REGION Network 3: Purga Bellis
   RUNG wire#powerrail
      Contact( "MC003" )
      Contact( "DB-PurgaComAlta".Habil_PurgaBellis )
      I_Contact( "Tag_55" )
      S_ODT(T_NO := "Tag_17", R := wire#w1, TV := #Aux1_MC003, BI =>, RET_VAL =>)
      wire#w2
      Coil( "MC003_EVP" )
   END_RUNG
   RUNG wire#powerrail
      I_Contact( "DB-PurgaComAlta".Habil_PurgaBellis )
   END_RUNG wire#w1
   RUNG wire#powerrail
      Contact( "DB-PurgaComAlta".Prueba_PurgaBellis )
      wire#w3
      I_Contact( "Tag_55" )
   END_RUNG wire#w2
   RUNG wire#powerrail
      Contact( "MC003_EVP" )
   END_RUNG wire#w3
   RUNG wire#w2
      S_ODT(T_NO := "Tag_55", TV := #Aux2_MC003, R :=, BI =>, RET_VAL =>)
   END_RUNG
   // the same network as SCL:
   #_s5time1 := S_ODT(T_NO := "Tag_17",
                      S := "MC003" AND "DB-PurgaComAlta".Habil_PurgaBellis AND NOT "Tag_55",
                      R := NOT "DB-PurgaComAlta".Habil_PurgaBellis,
                      TV := #Aux1_MC003,
                      Q => #_w1);
   "MC003_EVP" := #_w1 OR (("DB-PurgaComAlta".Prueba_PurgaBellis OR "MC003_EVP") AND NOT "Tag_55");
   #_s5time2 := S_ODT(T_NO := "Tag_55", S := "MC003_EVP", TV := #Aux2_MC003);
END_REGION

REGION Network 4
   RUNG wire#powerrail
      { S7_Templates := "SrcType := Int"; S7_GenerateENO := "TRUE" } Mul(in1 := "DB-PurgaComAlta".Toff_PurgaABC2, in2 := 6, out => #Aux1_MC001)
      { S7_Templates := "[SrcType := Int, DestType := Bcd16]"; S7_GenerateENO := "TRUE" } Convert(in := #Aux1_MC001, out => #Aux1_MC001)
      { S7_Templates := "SrcType := Int"; S7_GenerateENO := "TRUE" } Add(in1 := #Aux1_MC001, in2 := 16#3000, out => #Aux1_MC001)
   END_RUNG
   // the same network as SCL:
   // ENO of a box is taken as its EN; it also drops when the box reports an error
   #Aux1_MC001 := "DB-PurgaComAlta".Toff_PurgaABC2 * 6;
   #Aux1_MC001 := INT_TO_BCD16(#Aux1_MC001);
   #Aux1_MC001 := #Aux1_MC001 + 16#3000;
END_REGION

REGION Network 5
   RUNG wire#powerrail
      { S7_Templates := "SrcType := Int"; S7_GenerateENO := "TRUE" } Mul(in1 := "DB-PurgaComAlta".Ton_PurgaABC2, in2 := 10, out => #Aux2_MC001)
      { S7_Templates := "[SrcType := Int, DestType := Bcd16]"; S7_GenerateENO := "TRUE" } Convert(in := #Aux2_MC001, out => #Aux2_MC001)
      { S7_Templates := "SrcType := Int"; S7_GenerateENO := "TRUE" } Add(in1 := #Aux2_MC001, in2 := 16#1000, out => #Aux2_MC001)
   END_RUNG
   // the same network as SCL:
   // ENO of a box is taken as its EN; it also drops when the box reports an error
   #Aux2_MC001 := "DB-PurgaComAlta".Ton_PurgaABC2 * 10;
   #Aux2_MC001 := INT_TO_BCD16(#Aux2_MC001);
   #Aux2_MC001 := #Aux2_MC001 + 16#1000;
END_REGION

REGION Network 6: Purga ABC2
   RUNG wire#powerrail
      Contact( "MC001" )
      Contact( "DB-PurgaComAlta".Habil_PurgaABC2 )
      I_Contact( "Tag_65" )
      S_ODT(T_NO := "Tag_64", R := wire#w1, TV := #Aux1_MC001, BI =>, RET_VAL =>)
      I_Contact( "MC003_EVP" )
      wire#w2
      Coil( "MC001_EVP" )
   END_RUNG
   RUNG wire#powerrail
      I_Contact( "DB-PurgaComAlta".Habil_PurgaABC2 )
   END_RUNG wire#w1
   RUNG wire#powerrail
      Contact( "DB-PurgaComAlta".Prueba_PurgaABC2 )
      wire#w3
      I_Contact( "Tag_65" )
   END_RUNG wire#w2
   RUNG wire#powerrail
      Contact( "MC001_EVP" )
   END_RUNG wire#w3
   RUNG wire#w2
      S_ODT(T_NO := "Tag_65", TV := #Aux2_MC001, R :=, BI =>, RET_VAL =>)
   END_RUNG
   // the same network as SCL:
   #_s5time1 := S_ODT(T_NO := "Tag_64",
                      S := "MC001" AND "DB-PurgaComAlta".Habil_PurgaABC2 AND NOT "Tag_65",
                      R := NOT "DB-PurgaComAlta".Habil_PurgaABC2,
                      TV := #Aux1_MC001,
                      Q => #_w1);
   "MC001_EVP" := (#_w1 AND NOT "MC003_EVP") OR (("DB-PurgaComAlta".Prueba_PurgaABC2 OR "MC001_EVP") AND NOT "Tag_65");
   #_s5time2 := S_ODT(T_NO := "Tag_65", S := "MC001_EVP", TV := #Aux2_MC001);
END_REGION

REGION Network 7
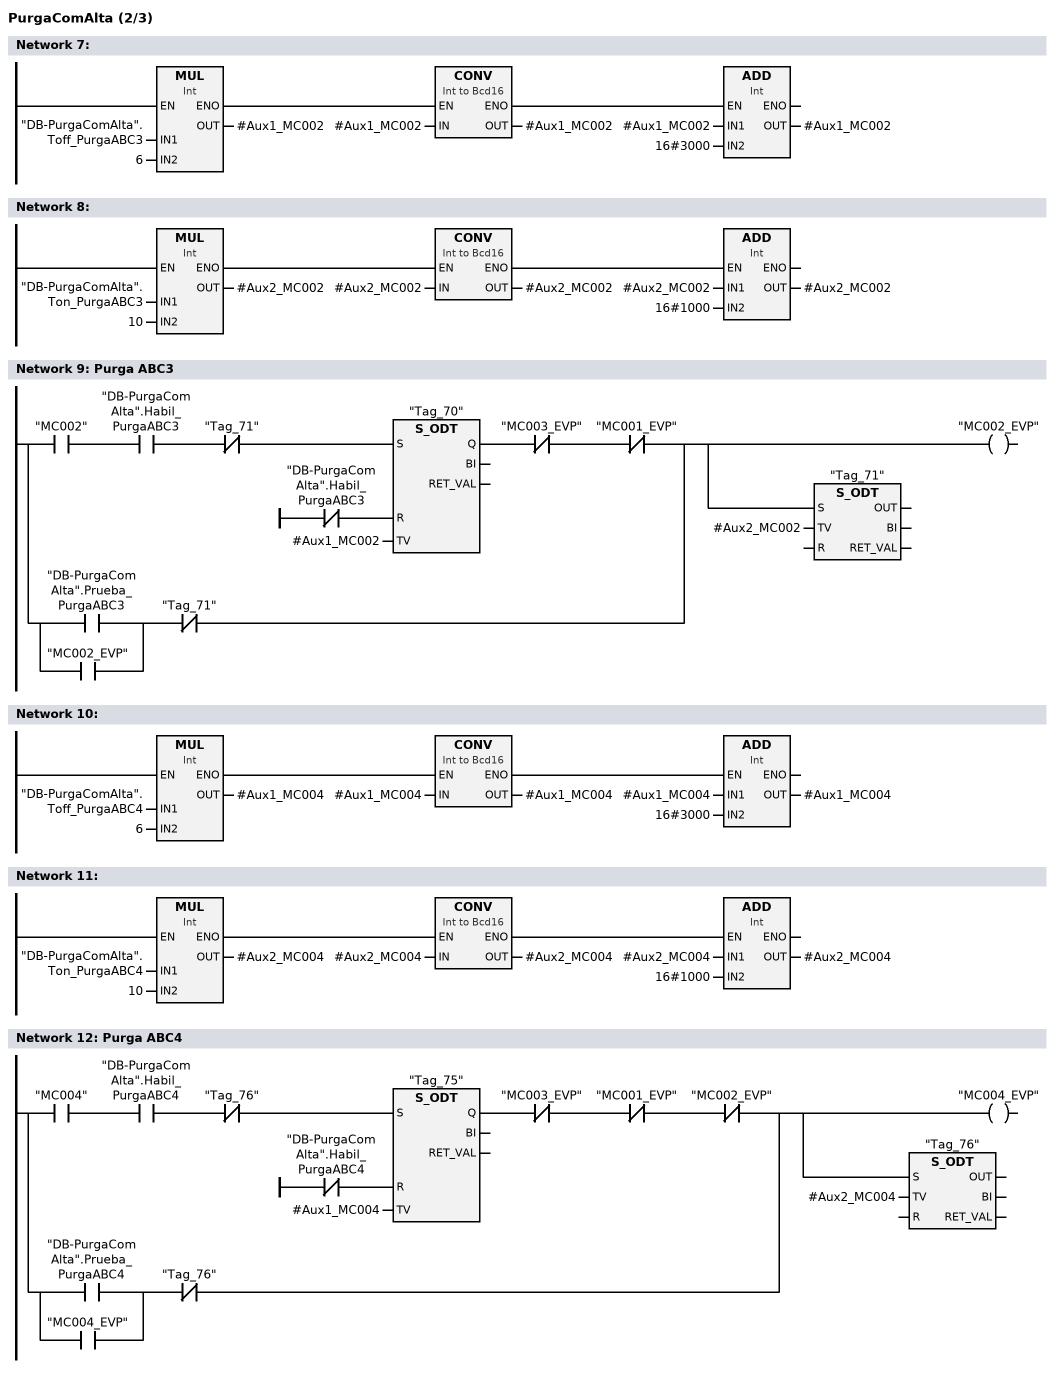
   RUNG wire#powerrail
      { S7_Templates := "SrcType := Int"; S7_GenerateENO := "TRUE" } Mul(in1 := "DB-PurgaComAlta".Toff_PurgaABC3, in2 := 6, out => #Aux1_MC002)
      { S7_Templates := "[SrcType := Int, DestType := Bcd16]"; S7_GenerateENO := "TRUE" } Convert(in := #Aux1_MC002, out => #Aux1_MC002)
      { S7_Templates := "SrcType := Int"; S7_GenerateENO := "TRUE" } Add(in1 := #Aux1_MC002, in2 := 16#3000, out => #Aux1_MC002)
   END_RUNG
   // the same network as SCL:
   // ENO of a box is taken as its EN; it also drops when the box reports an error
   #Aux1_MC002 := "DB-PurgaComAlta".Toff_PurgaABC3 * 6;
   #Aux1_MC002 := INT_TO_BCD16(#Aux1_MC002);
   #Aux1_MC002 := #Aux1_MC002 + 16#3000;
END_REGION

REGION Network 8
   RUNG wire#powerrail
      { S7_Templates := "SrcType := Int"; S7_GenerateENO := "TRUE" } Mul(in1 := "DB-PurgaComAlta".Ton_PurgaABC3, in2 := 10, out => #Aux2_MC002)
      { S7_Templates := "[SrcType := Int, DestType := Bcd16]"; S7_GenerateENO := "TRUE" } Convert(in := #Aux2_MC002, out => #Aux2_MC002)
      { S7_Templates := "SrcType := Int"; S7_GenerateENO := "TRUE" } Add(in1 := #Aux2_MC002, in2 := 16#1000, out => #Aux2_MC002)
   END_RUNG
   // the same network as SCL:
   // ENO of a box is taken as its EN; it also drops when the box reports an error
   #Aux2_MC002 := "DB-PurgaComAlta".Ton_PurgaABC3 * 10;
   #Aux2_MC002 := INT_TO_BCD16(#Aux2_MC002);
   #Aux2_MC002 := #Aux2_MC002 + 16#1000;
END_REGION

REGION Network 9: Purga ABC3
   RUNG wire#powerrail
      Contact( "MC002" )
      Contact( "DB-PurgaComAlta".Habil_PurgaABC3 )
      I_Contact( "Tag_71" )
      S_ODT(T_NO := "Tag_70", R := wire#w1, TV := #Aux1_MC002, BI =>, RET_VAL =>)
      I_Contact( "MC003_EVP" )
      I_Contact( "MC001_EVP" )
      wire#w2
      Coil( "MC002_EVP" )
   END_RUNG
   RUNG wire#powerrail
      I_Contact( "DB-PurgaComAlta".Habil_PurgaABC3 )
   END_RUNG wire#w1
   RUNG wire#powerrail
      Contact( "DB-PurgaComAlta".Prueba_PurgaABC3 )
      wire#w3
      I_Contact( "Tag_71" )
   END_RUNG wire#w2
   RUNG wire#powerrail
      Contact( "MC002_EVP" )
   END_RUNG wire#w3
   RUNG wire#w2
      S_ODT(T_NO := "Tag_71", TV := #Aux2_MC002, R :=, BI =>, RET_VAL =>)
   END_RUNG
   // the same network as SCL:
   #_s5time1 := S_ODT(T_NO := "Tag_70",
                      S := "MC002" AND "DB-PurgaComAlta".Habil_PurgaABC3 AND NOT "Tag_71",
                      R := NOT "DB-PurgaComAlta".Habil_PurgaABC3,
                      TV := #Aux1_MC002,
                      Q => #_w1);
   "MC002_EVP" := (#_w1 AND NOT "MC003_EVP" AND NOT "MC001_EVP") OR (("DB-PurgaComAlta".Prueba_PurgaABC3 OR "MC002_EVP") AND NOT "Tag_71");
   #_s5time2 := S_ODT(T_NO := "Tag_71", S := "MC002_EVP", TV := #Aux2_MC002);
END_REGION

REGION Network 10
   RUNG wire#powerrail
      { S7_Templates := "SrcType := Int"; S7_GenerateENO := "TRUE" } Mul(in1 := "DB-PurgaComAlta".Toff_PurgaABC4, in2 := 6, out => #Aux1_MC004)
      { S7_Templates := "[SrcType := Int, DestType := Bcd16]"; S7_GenerateENO := "TRUE" } Convert(in := #Aux1_MC004, out => #Aux1_MC004)
      { S7_Templates := "SrcType := Int"; S7_GenerateENO := "TRUE" } Add(in1 := #Aux1_MC004, in2 := 16#3000, out => #Aux1_MC004)
   END_RUNG
   // the same network as SCL:
   // ENO of a box is taken as its EN; it also drops when the box reports an error
   #Aux1_MC004 := "DB-PurgaComAlta".Toff_PurgaABC4 * 6;
   #Aux1_MC004 := INT_TO_BCD16(#Aux1_MC004);
   #Aux1_MC004 := #Aux1_MC004 + 16#3000;
END_REGION

REGION Network 11
   RUNG wire#powerrail
      { S7_Templates := "SrcType := Int"; S7_GenerateENO := "TRUE" } Mul(in1 := "DB-PurgaComAlta".Ton_PurgaABC4, in2 := 10, out => #Aux2_MC004)
      { S7_Templates := "[SrcType := Int, DestType := Bcd16]"; S7_GenerateENO := "TRUE" } Convert(in := #Aux2_MC004, out => #Aux2_MC004)
      { S7_Templates := "SrcType := Int"; S7_GenerateENO := "TRUE" } Add(in1 := #Aux2_MC004, in2 := 16#1000, out => #Aux2_MC004)
   END_RUNG
   // the same network as SCL:
   // ENO of a box is taken as its EN; it also drops when the box reports an error
   #Aux2_MC004 := "DB-PurgaComAlta".Ton_PurgaABC4 * 10;
   #Aux2_MC004 := INT_TO_BCD16(#Aux2_MC004);
   #Aux2_MC004 := #Aux2_MC004 + 16#1000;
END_REGION

REGION Network 12: Purga ABC4
   RUNG wire#powerrail
      Contact( "MC004" )
      Contact( "DB-PurgaComAlta".Habil_PurgaABC4 )
      I_Contact( "Tag_76" )
      S_ODT(T_NO := "Tag_75", R := wire#w1, TV := #Aux1_MC004, BI =>, RET_VAL =>)
      I_Contact( "MC003_EVP" )
      I_Contact( "MC001_EVP" )
      I_Contact( "MC002_EVP" )
      wire#w2
      Coil( "MC004_EVP" )
   END_RUNG
   RUNG wire#powerrail
      I_Contact( "DB-PurgaComAlta".Habil_PurgaABC4 )
   END_RUNG wire#w1
   RUNG wire#powerrail
      Contact( "DB-PurgaComAlta".Prueba_PurgaABC4 )
      wire#w3
      I_Contact( "Tag_76" )
   END_RUNG wire#w2
   RUNG wire#powerrail
      Contact( "MC004_EVP" )
   END_RUNG wire#w3
   RUNG wire#w2
      S_ODT(T_NO := "Tag_76", TV := #Aux2_MC004, R :=, BI =>, RET_VAL =>)
   END_RUNG
   // the same network as SCL:
   #_s5time1 := S_ODT(T_NO := "Tag_75",
                      S := "MC004" AND "DB-PurgaComAlta".Habil_PurgaABC4 AND NOT "Tag_76",
                      R := NOT "DB-PurgaComAlta".Habil_PurgaABC4,
                      TV := #Aux1_MC004,
                      Q => #_w1);
   "MC004_EVP" := (#_w1 AND NOT "MC003_EVP" AND NOT "MC001_EVP" AND NOT "MC002_EVP") OR (("DB-PurgaComAlta".Prueba_PurgaABC4 OR "MC004_EVP") AND NOT "Tag_76");
   #_s5time2 := S_ODT(T_NO := "Tag_76", S := "MC004_EVP", TV := #Aux2_MC004);
END_REGION

REGION Network 13
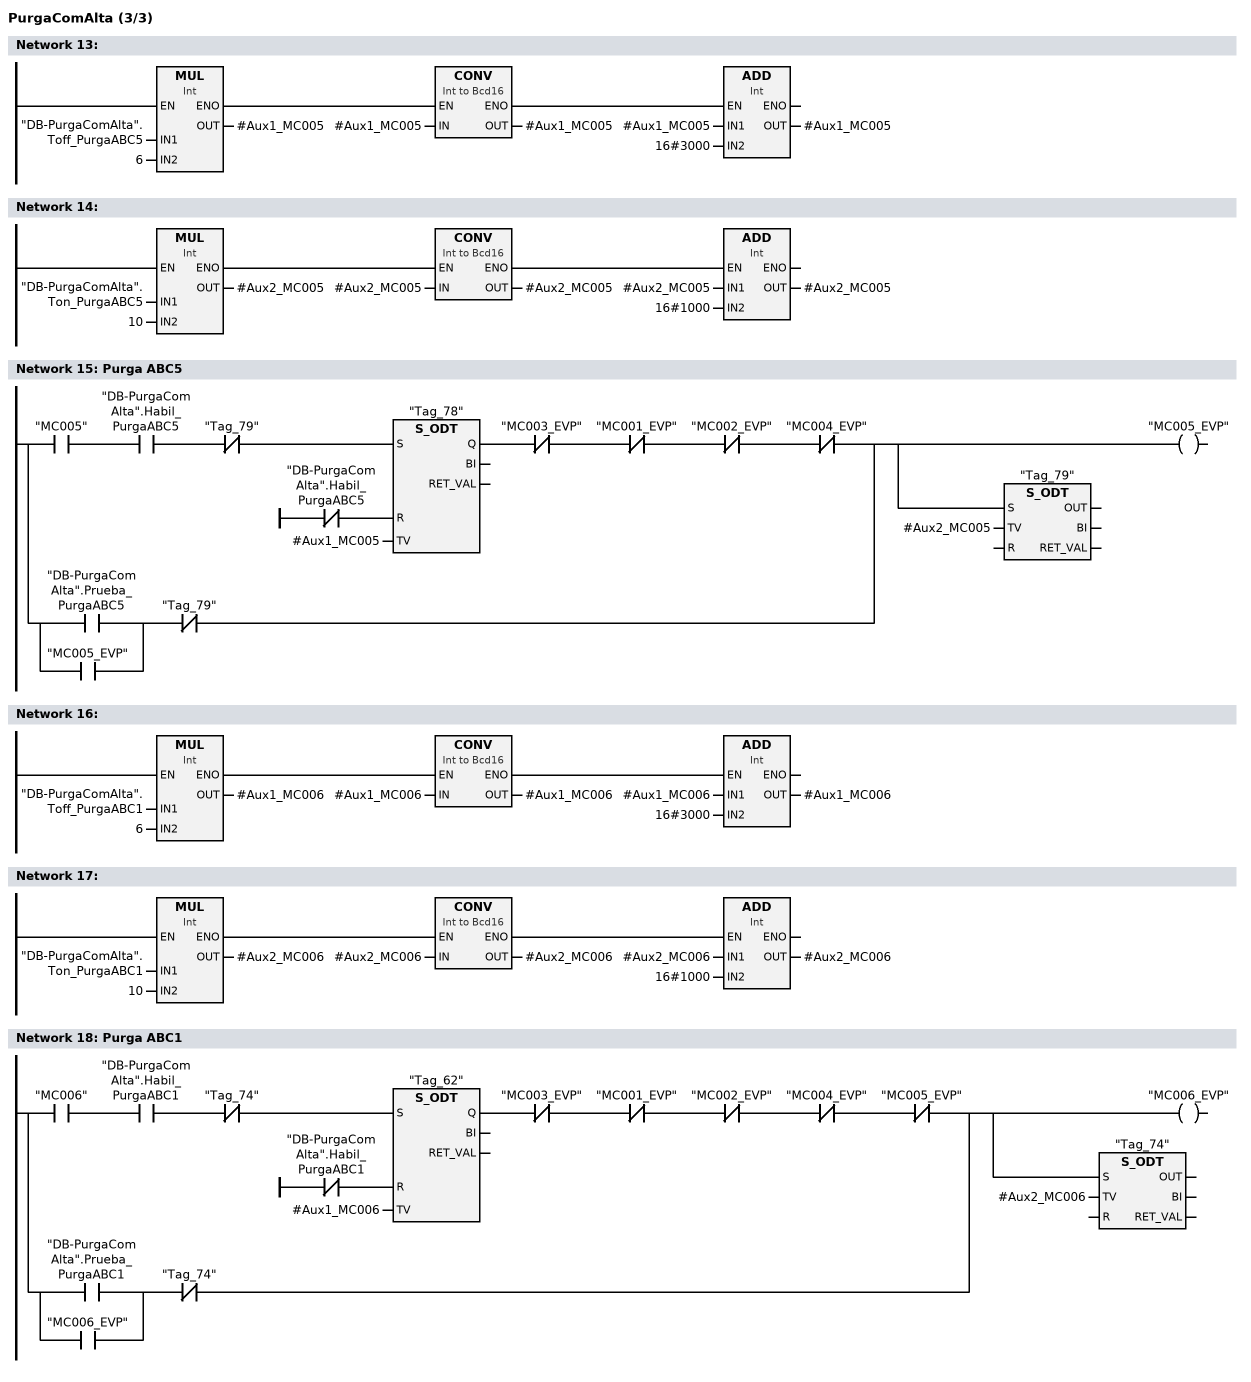
   RUNG wire#powerrail
      { S7_Templates := "SrcType := Int"; S7_GenerateENO := "TRUE" } Mul(in1 := "DB-PurgaComAlta".Toff_PurgaABC5, in2 := 6, out => #Aux1_MC005)
      { S7_Templates := "[SrcType := Int, DestType := Bcd16]"; S7_GenerateENO := "TRUE" } Convert(in := #Aux1_MC005, out => #Aux1_MC005)
      { S7_Templates := "SrcType := Int"; S7_GenerateENO := "TRUE" } Add(in1 := #Aux1_MC005, in2 := 16#3000, out => #Aux1_MC005)
   END_RUNG
   // the same network as SCL:
   // ENO of a box is taken as its EN; it also drops when the box reports an error
   #Aux1_MC005 := "DB-PurgaComAlta".Toff_PurgaABC5 * 6;
   #Aux1_MC005 := INT_TO_BCD16(#Aux1_MC005);
   #Aux1_MC005 := #Aux1_MC005 + 16#3000;
END_REGION

REGION Network 14
   RUNG wire#powerrail
      { S7_Templates := "SrcType := Int"; S7_GenerateENO := "TRUE" } Mul(in1 := "DB-PurgaComAlta".Ton_PurgaABC5, in2 := 10, out => #Aux2_MC005)
      { S7_Templates := "[SrcType := Int, DestType := Bcd16]"; S7_GenerateENO := "TRUE" } Convert(in := #Aux2_MC005, out => #Aux2_MC005)
      { S7_Templates := "SrcType := Int"; S7_GenerateENO := "TRUE" } Add(in1 := #Aux2_MC005, in2 := 16#1000, out => #Aux2_MC005)
   END_RUNG
   // the same network as SCL:
   // ENO of a box is taken as its EN; it also drops when the box reports an error
   #Aux2_MC005 := "DB-PurgaComAlta".Ton_PurgaABC5 * 10;
   #Aux2_MC005 := INT_TO_BCD16(#Aux2_MC005);
   #Aux2_MC005 := #Aux2_MC005 + 16#1000;
END_REGION

REGION Network 15: Purga ABC5
   RUNG wire#powerrail
      Contact( "MC005" )
      Contact( "DB-PurgaComAlta".Habil_PurgaABC5 )
      I_Contact( "Tag_79" )
      S_ODT(T_NO := "Tag_78", R := wire#w1, TV := #Aux1_MC005, BI =>, RET_VAL =>)
      I_Contact( "MC003_EVP" )
      I_Contact( "MC001_EVP" )
      I_Contact( "MC002_EVP" )
      I_Contact( "MC004_EVP" )
      wire#w2
      Coil( "MC005_EVP" )
   END_RUNG
   RUNG wire#powerrail
      I_Contact( "DB-PurgaComAlta".Habil_PurgaABC5 )
   END_RUNG wire#w1
   RUNG wire#powerrail
      Contact( "DB-PurgaComAlta".Prueba_PurgaABC5 )
      wire#w3
      I_Contact( "Tag_79" )
   END_RUNG wire#w2
   RUNG wire#powerrail
      Contact( "MC005_EVP" )
   END_RUNG wire#w3
   RUNG wire#w2
      S_ODT(T_NO := "Tag_79", TV := #Aux2_MC005, R :=, BI =>, RET_VAL =>)
   END_RUNG
   // the same network as SCL:
   #_s5time1 := S_ODT(T_NO := "Tag_78",
                      S := "MC005" AND "DB-PurgaComAlta".Habil_PurgaABC5 AND NOT "Tag_79",
                      R := NOT "DB-PurgaComAlta".Habil_PurgaABC5,
                      TV := #Aux1_MC005,
                      Q => #_w1);
   "MC005_EVP" := (#_w1 AND NOT "MC003_EVP" AND NOT "MC001_EVP" AND NOT "MC002_EVP" AND NOT "MC004_EVP") OR (("DB-PurgaComAlta".Prueba_PurgaABC5 OR "MC005_EVP") AND NOT "Tag_79");
   #_s5time2 := S_ODT(T_NO := "Tag_79", S := "MC005_EVP", TV := #Aux2_MC005);
END_REGION

REGION Network 16
   RUNG wire#powerrail
      { S7_Templates := "SrcType := Int"; S7_GenerateENO := "TRUE" } Mul(in1 := "DB-PurgaComAlta".Toff_PurgaABC1, in2 := 6, out => #Aux1_MC006)
      { S7_Templates := "[SrcType := Int, DestType := Bcd16]"; S7_GenerateENO := "TRUE" } Convert(in := #Aux1_MC006, out => #Aux1_MC006)
      { S7_Templates := "SrcType := Int"; S7_GenerateENO := "TRUE" } Add(in1 := #Aux1_MC006, in2 := 16#3000, out => #Aux1_MC006)
   END_RUNG
   // the same network as SCL:
   // ENO of a box is taken as its EN; it also drops when the box reports an error
   #Aux1_MC006 := "DB-PurgaComAlta".Toff_PurgaABC1 * 6;
   #Aux1_MC006 := INT_TO_BCD16(#Aux1_MC006);
   #Aux1_MC006 := #Aux1_MC006 + 16#3000;
END_REGION

REGION Network 17
   RUNG wire#powerrail
      { S7_Templates := "SrcType := Int"; S7_GenerateENO := "TRUE" } Mul(in1 := "DB-PurgaComAlta".Ton_PurgaABC1, in2 := 10, out => #Aux2_MC006)
      { S7_Templates := "[SrcType := Int, DestType := Bcd16]"; S7_GenerateENO := "TRUE" } Convert(in := #Aux2_MC006, out => #Aux2_MC006)
      { S7_Templates := "SrcType := Int"; S7_GenerateENO := "TRUE" } Add(in1 := #Aux2_MC006, in2 := 16#1000, out => #Aux2_MC006)
   END_RUNG
   // the same network as SCL:
   // ENO of a box is taken as its EN; it also drops when the box reports an error
   #Aux2_MC006 := "DB-PurgaComAlta".Ton_PurgaABC1 * 10;
   #Aux2_MC006 := INT_TO_BCD16(#Aux2_MC006);
   #Aux2_MC006 := #Aux2_MC006 + 16#1000;
END_REGION

REGION Network 18: Purga ABC1
   RUNG wire#powerrail
      Contact( "MC006" )
      Contact( "DB-PurgaComAlta".Habil_PurgaABC1 )
      I_Contact( "Tag_74" )
      S_ODT(T_NO := "Tag_62", R := wire#w1, TV := #Aux1_MC006, BI =>, RET_VAL =>)
      I_Contact( "MC003_EVP" )
      I_Contact( "MC001_EVP" )
      I_Contact( "MC002_EVP" )
      I_Contact( "MC004_EVP" )
      I_Contact( "MC005_EVP" )
      wire#w2
      Coil( "MC006_EVP" )
   END_RUNG
   RUNG wire#powerrail
      I_Contact( "DB-PurgaComAlta".Habil_PurgaABC1 )
   END_RUNG wire#w1
   RUNG wire#powerrail
      Contact( "DB-PurgaComAlta".Prueba_PurgaABC1 )
      wire#w3
      I_Contact( "Tag_74" )
   END_RUNG wire#w2
   RUNG wire#powerrail
      Contact( "MC006_EVP" )
   END_RUNG wire#w3
   RUNG wire#w2
      S_ODT(T_NO := "Tag_74", TV := #Aux2_MC006, R :=, BI =>, RET_VAL =>)
   END_RUNG
   // the same network as SCL:
   #_s5time1 := S_ODT(T_NO := "Tag_62",
                      S := "MC006" AND "DB-PurgaComAlta".Habil_PurgaABC1 AND NOT "Tag_74",
                      R := NOT "DB-PurgaComAlta".Habil_PurgaABC1,
                      TV := #Aux1_MC006,
                      Q => #_w1);
   "MC006_EVP" := (#_w1 AND NOT "MC003_EVP" AND NOT "MC001_EVP" AND NOT "MC002_EVP" AND NOT "MC004_EVP" AND NOT "MC005_EVP") OR (("DB-PurgaComAlta".Prueba_PurgaABC1 OR "MC006_EVP") AND NOT "Tag_74");
   #_s5time2 := S_ODT(T_NO := "Tag_74", S := "MC006_EVP", TV := #Aux2_MC006);
END_REGION
END_FUNCTION

// folder: Compresores/Alta/Máquina de Estados

FUNCTION "LogMaqEstGeneral" : Void   // FC35, LAD
{ S7_Optimized_Access := 'FALSE' }
VERSION : 0.1
   VAR_TEMP
      Temp_0 : Bool;
      Temp_1 : Bool;
      Temp_2 : Bool;
      Temp_3 : Bool;
      Temp_4 : Bool;
      Temp_5 : Bool;
      Temp_6 : Bool;
      Temp_7 : Bool;
      Temp_8 : Bool;
      Temp_9 : Bool;
      Temp_10 : Bool;
      Temp_11 : Bool;
   END_VAR
BEGIN

REGION Network 1
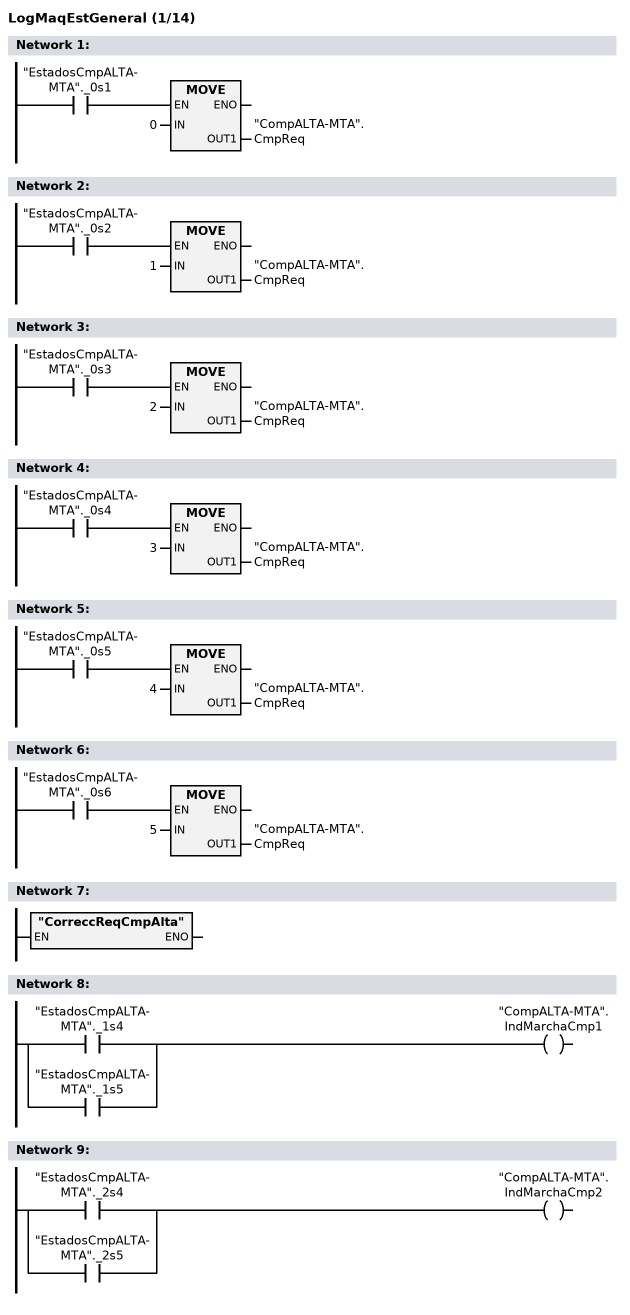
   RUNG wire#powerrail
      Contact( "EstadosCmpALTA-MTA"._0s1 )
      { S7_GenerateENO := "TRUE" } Move(in := 0, out1 => "CompALTA-MTA".CmpReq)
   END_RUNG
   // the same network as SCL:
   IF "EstadosCmpALTA-MTA"._0s1 THEN "CompALTA-MTA".CmpReq := 0; END_IF;
END_REGION

REGION Network 2
   RUNG wire#powerrail
      Contact( "EstadosCmpALTA-MTA"._0s2 )
      { S7_GenerateENO := "TRUE" } Move(in := 1, out1 => "CompALTA-MTA".CmpReq)
   END_RUNG
   // the same network as SCL:
   IF "EstadosCmpALTA-MTA"._0s2 THEN "CompALTA-MTA".CmpReq := 1; END_IF;
END_REGION

REGION Network 3
   RUNG wire#powerrail
      Contact( "EstadosCmpALTA-MTA"._0s3 )
      { S7_GenerateENO := "TRUE" } Move(in := 2, out1 => "CompALTA-MTA".CmpReq)
   END_RUNG
   // the same network as SCL:
   IF "EstadosCmpALTA-MTA"._0s3 THEN "CompALTA-MTA".CmpReq := 2; END_IF;
END_REGION

REGION Network 4
   RUNG wire#powerrail
      Contact( "EstadosCmpALTA-MTA"._0s4 )
      { S7_GenerateENO := "TRUE" } Move(in := 3, out1 => "CompALTA-MTA".CmpReq)
   END_RUNG
   // the same network as SCL:
   IF "EstadosCmpALTA-MTA"._0s4 THEN "CompALTA-MTA".CmpReq := 3; END_IF;
END_REGION

REGION Network 5
   RUNG wire#powerrail
      Contact( "EstadosCmpALTA-MTA"._0s5 )
      { S7_GenerateENO := "TRUE" } Move(in := 4, out1 => "CompALTA-MTA".CmpReq)
   END_RUNG
   // the same network as SCL:
   IF "EstadosCmpALTA-MTA"._0s5 THEN "CompALTA-MTA".CmpReq := 4; END_IF;
END_REGION

REGION Network 6
   RUNG wire#powerrail
      Contact( "EstadosCmpALTA-MTA"._0s6 )
      { S7_GenerateENO := "TRUE" } Move(in := 5, out1 => "CompALTA-MTA".CmpReq)
   END_RUNG
   // the same network as SCL:
   IF "EstadosCmpALTA-MTA"._0s6 THEN "CompALTA-MTA".CmpReq := 5; END_IF;
END_REGION

REGION Network 7
   RUNG wire#powerrail
      "CorreccReqCmpAlta"()
   END_RUNG
   // the same network as SCL:
   "CorreccReqCmpAlta"();
END_REGION

REGION Network 8
   RUNG wire#powerrail
      Contact( "EstadosCmpALTA-MTA"._1s4 )
      wire#w1
      Coil( "CompALTA-MTA".IndMarchaCmp1 )
   END_RUNG
   RUNG wire#powerrail
      Contact( "EstadosCmpALTA-MTA"._1s5 )
   END_RUNG wire#w1
   // the same network as SCL:
   "CompALTA-MTA".IndMarchaCmp1 := "EstadosCmpALTA-MTA"._1s4 OR "EstadosCmpALTA-MTA"._1s5;
END_REGION

REGION Network 9
   RUNG wire#powerrail
      Contact( "EstadosCmpALTA-MTA"._2s4 )
      wire#w1
      Coil( "CompALTA-MTA".IndMarchaCmp2 )
   END_RUNG
   RUNG wire#powerrail
      Contact( "EstadosCmpALTA-MTA"._2s5 )
   END_RUNG wire#w1
   // the same network as SCL:
   "CompALTA-MTA".IndMarchaCmp2 := "EstadosCmpALTA-MTA"._2s4 OR "EstadosCmpALTA-MTA"._2s5;
END_REGION

REGION Network 10
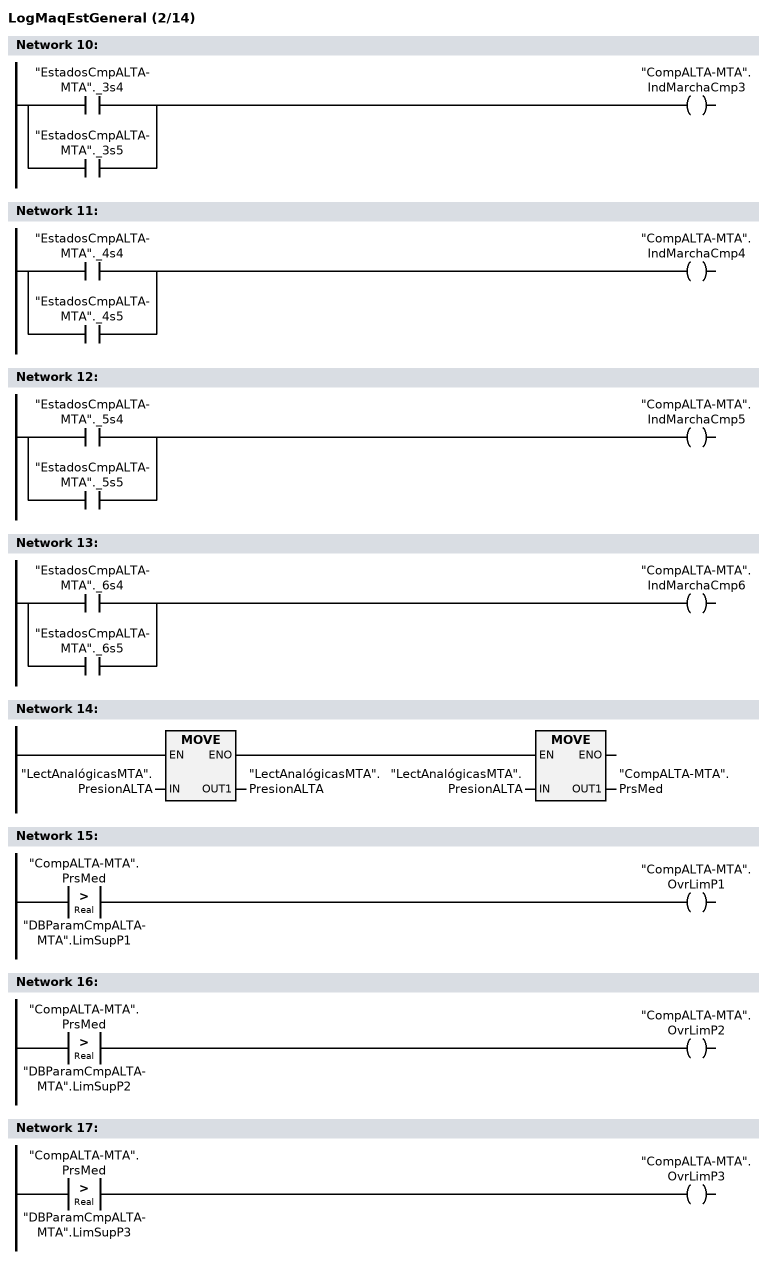
   RUNG wire#powerrail
      Contact( "EstadosCmpALTA-MTA"._3s4 )
      wire#w1
      Coil( "CompALTA-MTA".IndMarchaCmp3 )
   END_RUNG
   RUNG wire#powerrail
      Contact( "EstadosCmpALTA-MTA"._3s5 )
   END_RUNG wire#w1
   // the same network as SCL:
   "CompALTA-MTA".IndMarchaCmp3 := "EstadosCmpALTA-MTA"._3s4 OR "EstadosCmpALTA-MTA"._3s5;
END_REGION

REGION Network 11
   RUNG wire#powerrail
      Contact( "EstadosCmpALTA-MTA"._4s4 )
      wire#w1
      Coil( "CompALTA-MTA".IndMarchaCmp4 )
   END_RUNG
   RUNG wire#powerrail
      Contact( "EstadosCmpALTA-MTA"._4s5 )
   END_RUNG wire#w1
   // the same network as SCL:
   "CompALTA-MTA".IndMarchaCmp4 := "EstadosCmpALTA-MTA"._4s4 OR "EstadosCmpALTA-MTA"._4s5;
END_REGION

REGION Network 12
   RUNG wire#powerrail
      Contact( "EstadosCmpALTA-MTA"._5s4 )
      wire#w1
      Coil( "CompALTA-MTA".IndMarchaCmp5 )
   END_RUNG
   RUNG wire#powerrail
      Contact( "EstadosCmpALTA-MTA"._5s5 )
   END_RUNG wire#w1
   // the same network as SCL:
   "CompALTA-MTA".IndMarchaCmp5 := "EstadosCmpALTA-MTA"._5s4 OR "EstadosCmpALTA-MTA"._5s5;
END_REGION

REGION Network 13
   RUNG wire#powerrail
      Contact( "EstadosCmpALTA-MTA"._6s4 )
      wire#w1
      Coil( "CompALTA-MTA".IndMarchaCmp6 )
   END_RUNG
   RUNG wire#powerrail
      Contact( "EstadosCmpALTA-MTA"._6s5 )
   END_RUNG wire#w1
   // the same network as SCL:
   "CompALTA-MTA".IndMarchaCmp6 := "EstadosCmpALTA-MTA"._6s4 OR "EstadosCmpALTA-MTA"._6s5;
END_REGION

REGION Network 14
   RUNG wire#powerrail
      { S7_GenerateENO := "TRUE" } Move(in := "LectAnalógicasMTA".PresionALTA, out1 => "LectAnalógicasMTA".PresionALTA)
      { S7_GenerateENO := "TRUE" } Move(in := "LectAnalógicasMTA".PresionALTA, out1 => "CompALTA-MTA".PrsMed)
   END_RUNG
   // the same network as SCL:
   // ENO of a box is taken as its EN; it also drops when the box reports an error
   "LectAnalógicasMTA".PresionALTA := "LectAnalógicasMTA".PresionALTA;
   "CompALTA-MTA".PrsMed := "LectAnalógicasMTA".PresionALTA;
END_REGION

REGION Network 15
   RUNG wire#powerrail
      { S7_Templates := "SrcType := Real" } GT_Contact(in1 := "CompALTA-MTA".PrsMed, in2 := "DBParamCmpALTA-MTA".LimSupP1)
      Coil( "CompALTA-MTA".OvrLimP1 )
   END_RUNG
   // the same network as SCL:
   "CompALTA-MTA".OvrLimP1 := "CompALTA-MTA".PrsMed > "DBParamCmpALTA-MTA".LimSupP1;
END_REGION

REGION Network 16
   RUNG wire#powerrail
      { S7_Templates := "SrcType := Real" } GT_Contact(in1 := "CompALTA-MTA".PrsMed, in2 := "DBParamCmpALTA-MTA".LimSupP2)
      Coil( "CompALTA-MTA".OvrLimP2 )
   END_RUNG
   // the same network as SCL:
   "CompALTA-MTA".OvrLimP2 := "CompALTA-MTA".PrsMed > "DBParamCmpALTA-MTA".LimSupP2;
END_REGION

REGION Network 17
   RUNG wire#powerrail
      { S7_Templates := "SrcType := Real" } GT_Contact(in1 := "CompALTA-MTA".PrsMed, in2 := "DBParamCmpALTA-MTA".LimSupP3)
      Coil( "CompALTA-MTA".OvrLimP3 )
   END_RUNG
   // the same network as SCL:
   "CompALTA-MTA".OvrLimP3 := "CompALTA-MTA".PrsMed > "DBParamCmpALTA-MTA".LimSupP3;
END_REGION

REGION Network 18
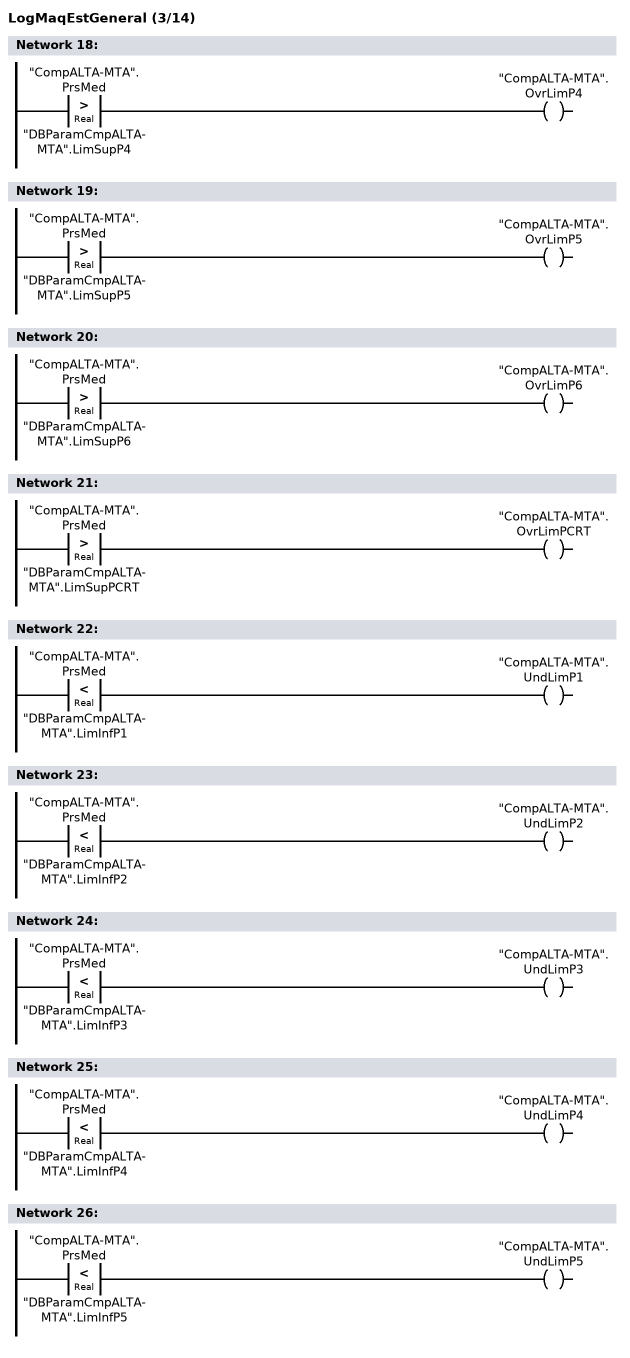
   RUNG wire#powerrail
      { S7_Templates := "SrcType := Real" } GT_Contact(in1 := "CompALTA-MTA".PrsMed, in2 := "DBParamCmpALTA-MTA".LimSupP4)
      Coil( "CompALTA-MTA".OvrLimP4 )
   END_RUNG
   // the same network as SCL:
   "CompALTA-MTA".OvrLimP4 := "CompALTA-MTA".PrsMed > "DBParamCmpALTA-MTA".LimSupP4;
END_REGION

REGION Network 19
   RUNG wire#powerrail
      { S7_Templates := "SrcType := Real" } GT_Contact(in1 := "CompALTA-MTA".PrsMed, in2 := "DBParamCmpALTA-MTA".LimSupP5)
      Coil( "CompALTA-MTA".OvrLimP5 )
   END_RUNG
   // the same network as SCL:
   "CompALTA-MTA".OvrLimP5 := "CompALTA-MTA".PrsMed > "DBParamCmpALTA-MTA".LimSupP5;
END_REGION

REGION Network 20
   RUNG wire#powerrail
      { S7_Templates := "SrcType := Real" } GT_Contact(in1 := "CompALTA-MTA".PrsMed, in2 := "DBParamCmpALTA-MTA".LimSupP6)
      Coil( "CompALTA-MTA".OvrLimP6 )
   END_RUNG
   // the same network as SCL:
   "CompALTA-MTA".OvrLimP6 := "CompALTA-MTA".PrsMed > "DBParamCmpALTA-MTA".LimSupP6;
END_REGION

REGION Network 21
   RUNG wire#powerrail
      { S7_Templates := "SrcType := Real" } GT_Contact(in1 := "CompALTA-MTA".PrsMed, in2 := "DBParamCmpALTA-MTA".LimSupPCRT)
      Coil( "CompALTA-MTA".OvrLimPCRT )
   END_RUNG
   // the same network as SCL:
   "CompALTA-MTA".OvrLimPCRT := "CompALTA-MTA".PrsMed > "DBParamCmpALTA-MTA".LimSupPCRT;
END_REGION

REGION Network 22
   RUNG wire#powerrail
      { S7_Templates := "SrcType := Real" } LT_Contact(in1 := "CompALTA-MTA".PrsMed, in2 := "DBParamCmpALTA-MTA".LimInfP1)
      Coil( "CompALTA-MTA".UndLimP1 )
   END_RUNG
   // the same network as SCL:
   "CompALTA-MTA".UndLimP1 := "CompALTA-MTA".PrsMed < "DBParamCmpALTA-MTA".LimInfP1;
END_REGION

REGION Network 23
   RUNG wire#powerrail
      { S7_Templates := "SrcType := Real" } LT_Contact(in1 := "CompALTA-MTA".PrsMed, in2 := "DBParamCmpALTA-MTA".LimInfP2)
      Coil( "CompALTA-MTA".UndLimP2 )
   END_RUNG
   // the same network as SCL:
   "CompALTA-MTA".UndLimP2 := "CompALTA-MTA".PrsMed < "DBParamCmpALTA-MTA".LimInfP2;
END_REGION

REGION Network 24
   RUNG wire#powerrail
      { S7_Templates := "SrcType := Real" } LT_Contact(in1 := "CompALTA-MTA".PrsMed, in2 := "DBParamCmpALTA-MTA".LimInfP3)
      Coil( "CompALTA-MTA".UndLimP3 )
   END_RUNG
   // the same network as SCL:
   "CompALTA-MTA".UndLimP3 := "CompALTA-MTA".PrsMed < "DBParamCmpALTA-MTA".LimInfP3;
END_REGION

REGION Network 25
   RUNG wire#powerrail
      { S7_Templates := "SrcType := Real" } LT_Contact(in1 := "CompALTA-MTA".PrsMed, in2 := "DBParamCmpALTA-MTA".LimInfP4)
      Coil( "CompALTA-MTA".UndLimP4 )
   END_RUNG
   // the same network as SCL:
   "CompALTA-MTA".UndLimP4 := "CompALTA-MTA".PrsMed < "DBParamCmpALTA-MTA".LimInfP4;
END_REGION

REGION Network 26
   RUNG wire#powerrail
      { S7_Templates := "SrcType := Real" } LT_Contact(in1 := "CompALTA-MTA".PrsMed, in2 := "DBParamCmpALTA-MTA".LimInfP5)
      Coil( "CompALTA-MTA".UndLimP5 )
   END_RUNG
   // the same network as SCL:
   "CompALTA-MTA".UndLimP5 := "CompALTA-MTA".PrsMed < "DBParamCmpALTA-MTA".LimInfP5;
END_REGION

REGION Network 27
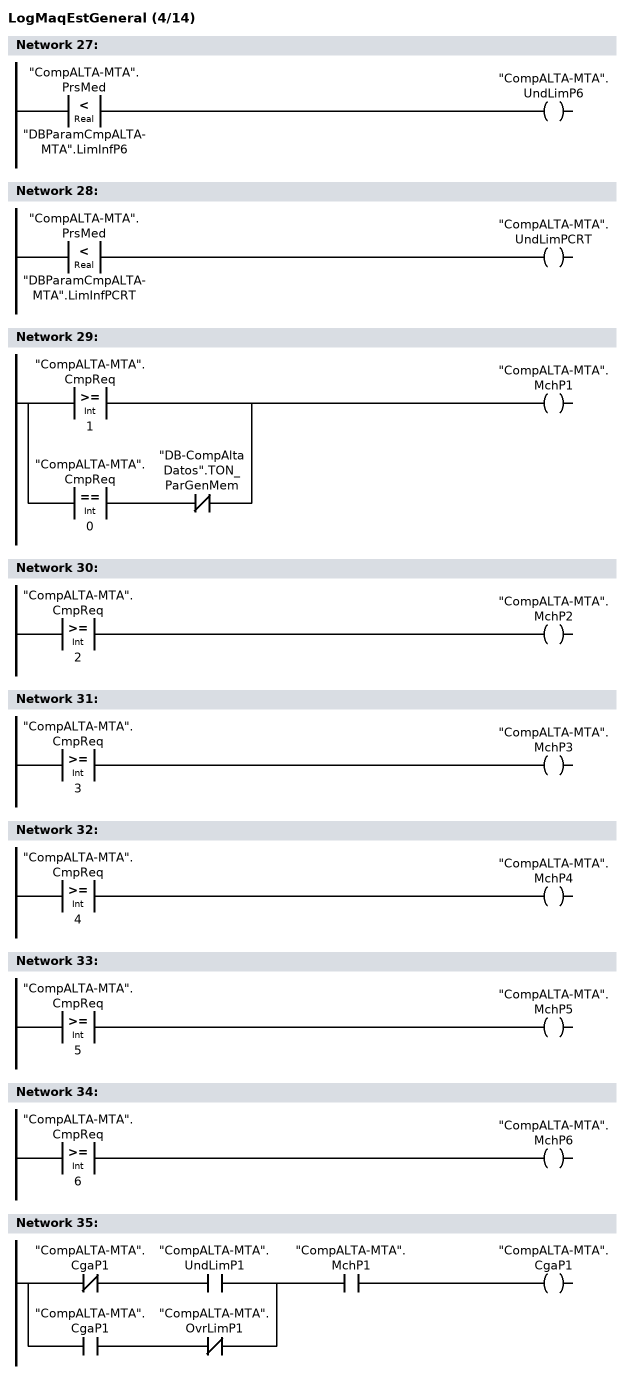
   RUNG wire#powerrail
      { S7_Templates := "SrcType := Real" } LT_Contact(in1 := "CompALTA-MTA".PrsMed, in2 := "DBParamCmpALTA-MTA".LimInfP6)
      Coil( "CompALTA-MTA".UndLimP6 )
   END_RUNG
   // the same network as SCL:
   "CompALTA-MTA".UndLimP6 := "CompALTA-MTA".PrsMed < "DBParamCmpALTA-MTA".LimInfP6;
END_REGION

REGION Network 28
   RUNG wire#powerrail
      { S7_Templates := "SrcType := Real" } LT_Contact(in1 := "CompALTA-MTA".PrsMed, in2 := "DBParamCmpALTA-MTA".LimInfPCRT)
      Coil( "CompALTA-MTA".UndLimPCRT )
   END_RUNG
   // the same network as SCL:
   "CompALTA-MTA".UndLimPCRT := "CompALTA-MTA".PrsMed < "DBParamCmpALTA-MTA".LimInfPCRT;
END_REGION

REGION Network 29
   RUNG wire#powerrail
      { S7_Templates := "SrcType := Int" } GE_Contact(in1 := "CompALTA-MTA".CmpReq, in2 := 1)
      wire#w1
      Coil( "CompALTA-MTA".MchP1 )
   END_RUNG
   RUNG wire#powerrail
      { S7_Templates := "SrcType := Int" } EQ_Contact(in1 := "CompALTA-MTA".CmpReq, in2 := 0)
      I_Contact( "DB-CompAltaDatos".TON_ParGenMem )
   END_RUNG wire#w1
   // the same network as SCL:
   "CompALTA-MTA".MchP1 := ("CompALTA-MTA".CmpReq >= 1) OR (("CompALTA-MTA".CmpReq = 0) AND NOT "DB-CompAltaDatos".TON_ParGenMem);
END_REGION

REGION Network 30
   RUNG wire#powerrail
      { S7_Templates := "SrcType := Int" } GE_Contact(in1 := "CompALTA-MTA".CmpReq, in2 := 2)
      Coil( "CompALTA-MTA".MchP2 )
   END_RUNG
   // the same network as SCL:
   "CompALTA-MTA".MchP2 := "CompALTA-MTA".CmpReq >= 2;
END_REGION

REGION Network 31
   RUNG wire#powerrail
      { S7_Templates := "SrcType := Int" } GE_Contact(in1 := "CompALTA-MTA".CmpReq, in2 := 3)
      Coil( "CompALTA-MTA".MchP3 )
   END_RUNG
   // the same network as SCL:
   "CompALTA-MTA".MchP3 := "CompALTA-MTA".CmpReq >= 3;
END_REGION

REGION Network 32
   RUNG wire#powerrail
      { S7_Templates := "SrcType := Int" } GE_Contact(in1 := "CompALTA-MTA".CmpReq, in2 := 4)
      Coil( "CompALTA-MTA".MchP4 )
   END_RUNG
   // the same network as SCL:
   "CompALTA-MTA".MchP4 := "CompALTA-MTA".CmpReq >= 4;
END_REGION

REGION Network 33
   RUNG wire#powerrail
      { S7_Templates := "SrcType := Int" } GE_Contact(in1 := "CompALTA-MTA".CmpReq, in2 := 5)
      Coil( "CompALTA-MTA".MchP5 )
   END_RUNG
   // the same network as SCL:
   "CompALTA-MTA".MchP5 := "CompALTA-MTA".CmpReq >= 5;
END_REGION

REGION Network 34
   RUNG wire#powerrail
      { S7_Templates := "SrcType := Int" } GE_Contact(in1 := "CompALTA-MTA".CmpReq, in2 := 6)
      Coil( "CompALTA-MTA".MchP6 )
   END_RUNG
   // the same network as SCL:
   "CompALTA-MTA".MchP6 := "CompALTA-MTA".CmpReq >= 6;
END_REGION

REGION Network 35
   RUNG wire#powerrail
      I_Contact( "CompALTA-MTA".CgaP1 )
      Contact( "CompALTA-MTA".UndLimP1 )
      wire#w1
      Contact( "CompALTA-MTA".MchP1 )
      Coil( "CompALTA-MTA".CgaP1 )
   END_RUNG
   RUNG wire#powerrail
      Contact( "CompALTA-MTA".CgaP1 )
      I_Contact( "CompALTA-MTA".OvrLimP1 )
   END_RUNG wire#w1
   // the same network as SCL:
   "CompALTA-MTA".CgaP1 := ((NOT "CompALTA-MTA".CgaP1 AND "CompALTA-MTA".UndLimP1) OR ("CompALTA-MTA".CgaP1 AND NOT "CompALTA-MTA".OvrLimP1)) AND "CompALTA-MTA".MchP1;
END_REGION

REGION Network 36
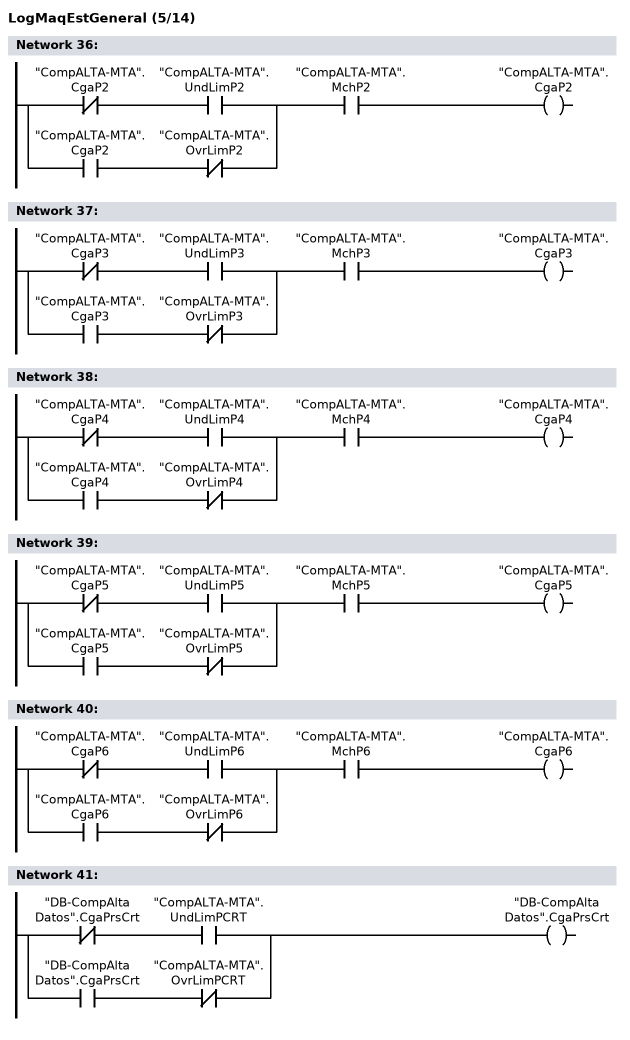
   RUNG wire#powerrail
      I_Contact( "CompALTA-MTA".CgaP2 )
      Contact( "CompALTA-MTA".UndLimP2 )
      wire#w1
      Contact( "CompALTA-MTA".MchP2 )
      Coil( "CompALTA-MTA".CgaP2 )
   END_RUNG
   RUNG wire#powerrail
      Contact( "CompALTA-MTA".CgaP2 )
      I_Contact( "CompALTA-MTA".OvrLimP2 )
   END_RUNG wire#w1
   // the same network as SCL:
   "CompALTA-MTA".CgaP2 := ((NOT "CompALTA-MTA".CgaP2 AND "CompALTA-MTA".UndLimP2) OR ("CompALTA-MTA".CgaP2 AND NOT "CompALTA-MTA".OvrLimP2)) AND "CompALTA-MTA".MchP2;
END_REGION

REGION Network 37
   RUNG wire#powerrail
      I_Contact( "CompALTA-MTA".CgaP3 )
      Contact( "CompALTA-MTA".UndLimP3 )
      wire#w1
      Contact( "CompALTA-MTA".MchP3 )
      Coil( "CompALTA-MTA".CgaP3 )
   END_RUNG
   RUNG wire#powerrail
      Contact( "CompALTA-MTA".CgaP3 )
      I_Contact( "CompALTA-MTA".OvrLimP3 )
   END_RUNG wire#w1
   // the same network as SCL:
   "CompALTA-MTA".CgaP3 := ((NOT "CompALTA-MTA".CgaP3 AND "CompALTA-MTA".UndLimP3) OR ("CompALTA-MTA".CgaP3 AND NOT "CompALTA-MTA".OvrLimP3)) AND "CompALTA-MTA".MchP3;
END_REGION

REGION Network 38
   RUNG wire#powerrail
      I_Contact( "CompALTA-MTA".CgaP4 )
      Contact( "CompALTA-MTA".UndLimP4 )
      wire#w1
      Contact( "CompALTA-MTA".MchP4 )
      Coil( "CompALTA-MTA".CgaP4 )
   END_RUNG
   RUNG wire#powerrail
      Contact( "CompALTA-MTA".CgaP4 )
      I_Contact( "CompALTA-MTA".OvrLimP4 )
   END_RUNG wire#w1
   // the same network as SCL:
   "CompALTA-MTA".CgaP4 := ((NOT "CompALTA-MTA".CgaP4 AND "CompALTA-MTA".UndLimP4) OR ("CompALTA-MTA".CgaP4 AND NOT "CompALTA-MTA".OvrLimP4)) AND "CompALTA-MTA".MchP4;
END_REGION

REGION Network 39
   RUNG wire#powerrail
      I_Contact( "CompALTA-MTA".CgaP5 )
      Contact( "CompALTA-MTA".UndLimP5 )
      wire#w1
      Contact( "CompALTA-MTA".MchP5 )
      Coil( "CompALTA-MTA".CgaP5 )
   END_RUNG
   RUNG wire#powerrail
      Contact( "CompALTA-MTA".CgaP5 )
      I_Contact( "CompALTA-MTA".OvrLimP5 )
   END_RUNG wire#w1
   // the same network as SCL:
   "CompALTA-MTA".CgaP5 := ((NOT "CompALTA-MTA".CgaP5 AND "CompALTA-MTA".UndLimP5) OR ("CompALTA-MTA".CgaP5 AND NOT "CompALTA-MTA".OvrLimP5)) AND "CompALTA-MTA".MchP5;
END_REGION

REGION Network 40
   RUNG wire#powerrail
      I_Contact( "CompALTA-MTA".CgaP6 )
      Contact( "CompALTA-MTA".UndLimP6 )
      wire#w1
      Contact( "CompALTA-MTA".MchP6 )
      Coil( "CompALTA-MTA".CgaP6 )
   END_RUNG
   RUNG wire#powerrail
      Contact( "CompALTA-MTA".CgaP6 )
      I_Contact( "CompALTA-MTA".OvrLimP6 )
   END_RUNG wire#w1
   // the same network as SCL:
   "CompALTA-MTA".CgaP6 := ((NOT "CompALTA-MTA".CgaP6 AND "CompALTA-MTA".UndLimP6) OR ("CompALTA-MTA".CgaP6 AND NOT "CompALTA-MTA".OvrLimP6)) AND "CompALTA-MTA".MchP6;
END_REGION

REGION Network 41
   RUNG wire#powerrail
      I_Contact( "DB-CompAltaDatos".CgaPrsCrt )
      Contact( "CompALTA-MTA".UndLimPCRT )
      wire#w1
      Coil( "DB-CompAltaDatos".CgaPrsCrt )
   END_RUNG
   RUNG wire#powerrail
      Contact( "DB-CompAltaDatos".CgaPrsCrt )
      I_Contact( "CompALTA-MTA".OvrLimPCRT )
   END_RUNG wire#w1
   // the same network as SCL:
   "DB-CompAltaDatos".CgaPrsCrt := (NOT "DB-CompAltaDatos".CgaPrsCrt AND "CompALTA-MTA".UndLimPCRT) OR ("DB-CompAltaDatos".CgaPrsCrt AND NOT "CompALTA-MTA".OvrLimPCRT);
END_REGION

REGION Network 42
